
                   // Segundo Convertir a DWORD y hacer SWAP para que el KRC lo lea correctamente
                   #moveCodeKuka := SWAP(UINT_TO_WORD(#code_int));
                   // "moveCodeKuka" := SWAP(UINT_TO_WORD(#code_int));

                   // Dispara GO (flanco por nivel)
                   "goTrigger" := NOT "goTrigger";     // Dispara pedido

                   // Marca estado/ack interno
                   #PlcStatusExecAccepted := TRUE;
                   #PlcStatusExecBusy := TRUE;
                   #PlcStatusExecDone := FALSE;

                   #lastSeq := #KukaControlCmdSeq;          // <-- memoriza!
                   #lastCode := #code_int;             // memoriza qué comando es (para actualizar activos en DONE)

                   #state := 20;                    // BUSY


       END_IF;

   20: // BUSY

       #PlcStatusExecBusy := TRUE;

       #code_int := #KukaControlCmdCode;

       // CANCEL pedido en BUSY → avisar al KRC y ACK de la ORDEN ACTIVA
       IF #code_int = 903 THEN
           "cancelGo" := TRUE;
       END_IF;

       IF ("rbDone" = "goTrigger") THEN
           // Fin confirmado por KUKA

           #PlcStatusExecDone := TRUE;
           #PlcStatusExecBusy := FALSE;
           #PlcStatusExecAccepted := FALSE;
           // ACK de la orden completada
           #PlcStatusExecAckSeq := #lastSeq;

           #state := 0;                         // vuelve a IDLE

       END_IF;

   30: // DONE
       // limpiar y volver a IDLE
       #state := 0;


   END_CASE;
END_REGION
END_FUNCTION_BLOCK

// folder: 20. Robot Services/RobotPos

FUNCTION_BLOCK "TcpPoseDecoderLe32"   // FB4, LAD
{ S7_Optimized_Access := 'TRUE' }
VERSION : 0.1
// Decodifica con SWAP, convierte a DINT y escala.
   VAR_INPUT
      xIniRawLe : DWord;
      yIniRawLe : DWord;
      zIniRawLe : DWord;
      e1IniRawLe : DWord;
      xFinRawLe : DWord;
      yFinRawLe : DWord;
      zFinRawLe : DWord;
      e1FinRawLe : DWord;
      ToolActiveRawByte : Byte;
      BaseActiveRawByte : Byte;
   END_VAR
   VAR_OUTPUT
      tcpPosIniX_mm : LReal;
      tcpPosIniY_mm : LReal;
      tcpPosIniZ_mm : LReal;
      e1PosIni_mm : LReal;
      tcpPosFinX_mm : LReal;
      tcpPosFinY_mm : LReal;
      tcpPosFinZ_mm : LReal;
      e1PosFin_mm : LReal;
      toolActiveId : UDInt;
      baseActiveId : UDInt;
   END_VAR
   VAR_TEMP
      xIniDint : DInt;
      yIniDint : DInt;
      zIniDint : DInt;
      aDint : DInt;
      bDint : DInt;
      cDint : DInt;
      e1IniDint : DInt;
      xFinDint : DInt;
      yFinDint : DInt;
      zFinDint : DInt;
      e1FinDint : DInt;
   END_VAR
BEGIN

REGION Network 1 (SCL): // 1) Endianness: ABCD -> DCBA
   #xIniDint := DWORD_TO_DINT(SWAP(#xIniRawLe));
   #yIniDint := DWORD_TO_DINT(SWAP(#yIniRawLe));
   #zIniDint := DWORD_TO_DINT(SWAP(#zIniRawLe));

   #e1IniDint := DWORD_TO_DINT(SWAP(#e1IniRawLe));

   #xFinDint := DWORD_TO_DINT(SWAP(#xFinRawLe));
   #yFinDint := DWORD_TO_DINT(SWAP(#yFinRawLe));
   #zFinDint := DWORD_TO_DINT(SWAP(#zFinRawLe));
   #e1FinDint := DWORD_TO_DINT(SWAP(#e1FinRawLe));
END_REGION

REGION Network 2 (SCL): // 2) Escala fixed-point: µm->mm, mdeg->deg
   #tcpPosIniX_mm := DINT_TO_LREAL(#xIniDint) / 1000.0;
   #tcpPosIniY_mm := DINT_TO_LREAL(#yIniDint) / 1000.0;
   #tcpPosIniZ_mm := DINT_TO_LREAL(#zIniDint) / 1000.0;

   #e1PosIni_mm := DINT_TO_LREAL(#e1IniDint) / 1000.0;  // mm o deg según tu E1

   #tcpPosFinX_mm := DINT_TO_LREAL(#xFinDint) / 1000.0;
   #tcpPosFinY_mm := DINT_TO_LREAL(#yFinDint) / 1000.0;
   #tcpPosFinZ_mm := DINT_TO_LREAL(#zFinDint) / 1000.0;
   #e1PosFin_mm := DINT_TO_LREAL(#e1FinDint) / 1000.0;  // mm o deg según tu E1

   #toolActiveId := #ToolActiveRawByte;
   #baseActiveId := #BaseActiveRawByte;
END_REGION
END_FUNCTION_BLOCK

// folder: 20. Robot Services/Tooling & Parking

FUNCTION_BLOCK "ToolChange"   // FB6, LAD
TITLE = FB: ManageTed009Station
{ S7_Optimized_Access := 'TRUE' }
VERSION : 0.1
// //  - KUKA manda órdenes (kukaCmd*)
// //  - El FB acciona bobinas de la docking (dockValve*On)
// //  - El FB publica ecos/estados para el KUKA (kukaFeedback*)
// //  - V2 (Unlock) puede mantenerse automática con útil aparcado
// //    (AutoUnlockWhenToolPresent = TRUE) [REF: estándar automático]. 
// //    Con útil ausente, no se activa para evitar soplado innecesario.
// //  - Tapa: FSM con interlock de zona segura y timeouts simétricos.
// //  - Diagnóstico: diagStep/diagFault/diagFaultCode.
// //
// //  Referencias (ver manual Stäubli TED009):
// //    • Sequence plan y sondeo ~20 ms durante conectar/desconectar. 
// //    • +21 mm: E2=0 ∧ E3=1 ∧ D1=0 antes de acoplar. 
// //    • z=0: bloquear retirando V2 y esperar E2=1 ∧ D1=1 (+E1=1). 
// //    • Retiradas +10/+70 y +25/>29 (comentadas para el programa del robot).
   VAR_INPUT
      kukaCmdOpenCover : Bool;
      kukaCmdCloseCover : Bool;
      kukaCmdUnlockMps : Bool;
      kukaCmdSafeForChange : Bool;
      dockSensorToolInPosition : Bool;   // E6
      dockSensorCoverClosed : Bool;   // E4
      dockSensorCoverOpen : Bool;   // E5
      robotSensorMpsUnlocked : Bool;   // E3
      robotSensorMpsLocked : Bool;   // E2
      robotSensorMpsCoupled : Bool;   // E1
      robotSensorMpsCtrlAirPressureOk : Bool;   // D1
      resetFault : Bool;
   END_VAR
   VAR_OUTPUT
      dockValveCoverOpenOn : Bool;   // bobina abrir tapa
      dockValveCoverCloseOn : Bool;   // bobina cerrar tapa
      dockValveV2UnlockOn : Bool;   // V2: aire de desbloqueo hacia módulo del robot
      MpsValveV1B12S4_ON : Bool;
      kukaFeedbackDockCoverOpen : Bool;
      kukaFeedbackDockCoverClosed : Bool;
      kukaFeedbackRobotMpsUnlocked : Bool;
      kukaFeedbackRobotMpsLocked : Bool;
      kukaFeedbackRobotMpsCoupled : Bool;
      kukaFeedbackMpsCtrlAirPressureOk : Bool;
      kukaFeedbackDockToolInPosition : Bool;
      diagStep : Int;
      diagFault : Bool;
      diagFaultCode : Int;
   END_VAR
   VAR
      "step" : Int;
      fault : Bool;
      faultCode : Int;
      AutoUnlockWhenToolPresent : Bool := true;   // // modo auto
      coverTimeout : Time := T#8S;   // // timeout de tapa (abrir/cerrar)
      unlockTimeout : Time := T#2S;   // // timeout de UNLOCK (E3=1 & D1=0)
      unlockReq : Bool;
      unlockReqEnabled : Bool;
      tempCoverOpen : TON_TIME;
      tempCoverClose : TON_TIME;
      tempUnlock : TON_TIME;
      autoUnlockEligible : Bool;
   END_VAR
   VAR CONSTANT
      StateIdle : Int := 0;
      StateOpening : Int := 10;
      StateOpen : Int := 11;
      StateClosing : Int := 20;
      StateClosed : Int := 21;
      FaultNone : Int;
      FaultOpenTimeout : Int := 101;
      FaultCloseTimeout : Int := 102;
      FaultUnlockTimeout : Int := 201;
      FaultInterlock : Int := 301;
   END_VAR
BEGIN

REGION Network 1 (SCL): Lógica de tapa + V2 (Unlock) de la docking
   // --- Feedbacks de estados al robot (eco directo de sensores físicos)
   #kukaFeedbackDockToolInPosition := #dockSensorToolInPosition; // E6 - herramienta en docking station
   #kukaFeedbackDockCoverOpen := #dockSensorCoverOpen;         // E4 - tapa abierta
   #kukaFeedbackDockCoverClosed := #dockSensorCoverClosed;     // E5 - tapa cerrada
   #kukaFeedbackRobotMpsUnlocked := #robotSensorMpsUnlocked;  // E3 - MPS desbloqueado (robot side)
   #kukaFeedbackRobotMpsLocked := #robotSensorMpsLocked;     // E2 - MPS bloqueado (robot side
   #kukaFeedbackRobotMpsCoupled := #robotSensorMpsCoupled;        // E1 - MPS acoplado  (robot side) 
   #kukaFeedbackMpsCtrlAirPressureOk := #robotSensorMpsCtrlAirPressureOk;  // D1 -presostato módulo aire control (robot)
   // ---- Reset de fallos/estado -------------------------------------------
   // Permite reconocer fallos desde HMI/Robot. Pone las salidas a 0 y la FSM (flow state machine)
   // Deja el FB en reposo (IDLE), corta bobinas y reinicia tempor TONs.
   // 
   IF #resetFault THEN
       #fault := FALSE;
       #faultCode := #FaultNone;
       #step := #StateIdle;

       #dockValveCoverOpenOn := FALSE;
       #dockValveCoverCloseOn := FALSE;
       #dockValveV2UnlockOn := FALSE;

       // Reset explícito de TON: IN=FALSE + PT definido
       #tempCoverOpen(IN := FALSE,
                      PT := #coverTimeout);
       #tempCoverClose(IN := FALSE,
                       PT := #coverTimeout);
       #tempUnlock(IN := FALSE,
                   PT := #unlockTimeout);
   END_IF;

   // ================= LÓGICA DE TAPA (máquina de estados) =================
   // Interlock básico: no se permite accionar tapa si el robot no confirma zona segura
   // (manual: abrir/cerrar solo fuera del barrido).
   CASE #step OF

       #StateIdle: // IDLE
           // Reposo ( tapa sin accionar); evaluar órdenes de KUKA.
           #dockValveCoverOpenOn := FALSE;
           #dockValveCoverCloseOn := FALSE;

           IF #kukaCmdSafeForChange THEN
               // Abrir si lo pide el robot y aún no está abierta
               IF (#kukaCmdOpenCover AND NOT #dockSensorCoverOpen) THEN
                   #step := #StateOpening;
               END_IF;
               // Cerrar si lo pide el robot y aún no está cerrada
               IF (#kukaCmdCloseCover AND NOT #dockSensorCoverClosed) THEN
                   #step := #StateClosing;
               END_IF;
           ELSIF (#kukaCmdOpenCover OR #kukaCmdCloseCover) THEN
               // Petición sin zona segura -> fallo de interlock
               #fault := TRUE;
               #faultCode := #FaultInterlock; // robot no garantiza zona segura
           END_IF;

       #StateOpening:  // Abrir tapa
           #dockValveCoverOpenOn := TRUE;
           #dockValveCoverCloseOn := FALSE;

           // Timeout de apertura: si no llega "tapa abierta" dentro de coverTimeout -> fallo.
           // coverTimeout debe ser > 3 s (tiempo típico de maniobra)
           #tempCoverOpen(IN := NOT #dockSensorCoverOpen,
                          PT := #coverTimeout);

           IF (#dockSensorCoverOpen AND NOT #dockSensorCoverClosed) THEN
               #tempCoverOpen(IN := FALSE,
                              PT := #coverTimeout);
               #step := #StateOpen;
           ELSIF #tempCoverOpen.Q THEN
               #fault := TRUE;
               #faultCode := #FaultOpenTimeout;
               #dockValveCoverOpenOn := FALSE;
               #step := #StateIdle;
           END_IF;

       #StateOpen: // Tapa abierta (estable)
           #dockValveCoverOpenOn := FALSE;
           #dockValveCoverCloseOn := FALSE;

           IF (#kukaCmdSafeForChange AND #kukaCmdCloseCover) THEN
               #step := #StateClosing;
           END_IF;


       #StateClosing: // Cerrar tapa
           #dockValveCoverOpenOn := FALSE;
           #dockValveCoverCloseOn := TRUE;

           // Timeout de cierre: si no llega "tapa cerrada" dentro de coverTimeout -> fallo.
           #tempCoverClose(IN := NOT #dockSensorCoverClosed,
                           PT := #coverTimeout);

           IF (#dockSensorCoverClosed AND NOT #dockSensorCoverOpen) THEN
               #tempCoverClose(IN := FALSE,
                               PT := #coverTimeout);
               #step := #StateClosed;
           ELSIF #tempCoverClose.Q THEN
               #fault := TRUE;
               #faultCode := #FaultCloseTimeout;
               #dockValveCoverCloseOn := FALSE;
               #step := #StateIdle;
           END_IF;

       #StateClosed: // Tapa cerrada (estable)
           #dockValveCoverOpenOn := FALSE;
           #dockValveCoverCloseOn := FALSE;

           IF (#kukaCmdSafeForChange AND #kukaCmdOpenCover) THEN
               #step := #StateOpening;
           END_IF;

       ELSE
           #step := #StateIdle;
   END_CASE;

   // Exclusión mutua de bobinas de tapa (seguridad por si alguna rama dejó ambas a 1)
   IF #dockValveCoverOpenOn THEN
       #dockValveCoverCloseOn := FALSE;
   END_IF;
   IF #dockValveCoverCloseOn THEN
       #dockValveCoverOpenOn := FALSE;
   END_IF;



   // -------- Arbitraje de V2 (UNLOCK) — sin auto-unlock --------
   #autoUnlockEligible := FALSE;   // DEPRECATED: ya no se usa

   //Cuando el robot va al punto de acople hace antes kukaCmdUnlockMpsYugo = TRUE

   //  solo por orden KUKA 
   #dockValveV2UnlockOn := #kukaCmdUnlockMps;

   IF #robotSensorMpsLocked THEN
       #MpsValveV1B12S4_ON := TRUE;
   END_IF;


   // Supervisión del estado desbloqueado (E3=1 y D1=0 en tiempo):
   #tempUnlock(
               IN := (#dockValveV2UnlockOn
               AND NOT (#robotSensorMpsUnlocked
               AND NOT #robotSensorMpsCtrlAirPressureOk)),
               PT := #unlockTimeout
   );
   IF NOT #dockValveV2UnlockOn THEN
       // reset explícito del TON cuando ya no se pide V2
       #tempUnlock(IN := FALSE,
                   PT := #unlockTimeout);
   END_IF;

   // -------------------- DIAGNÓSTICO PUBLICADO ----------------------------
   #diagStep := #step; // StateIdle/Opening/Open/Closing/Closed
   #diagFault := #fault;
   #diagFaultCode := #faultCode;
END_REGION
END_FUNCTION_BLOCK

FUNCTION_BLOCK "MpsDockingStation"   // FB9, LAD
{ S7_Optimized_Access := 'TRUE' }
VERSION : 0.1
BEGIN

REGION Network 1: Identificador de Herramienta
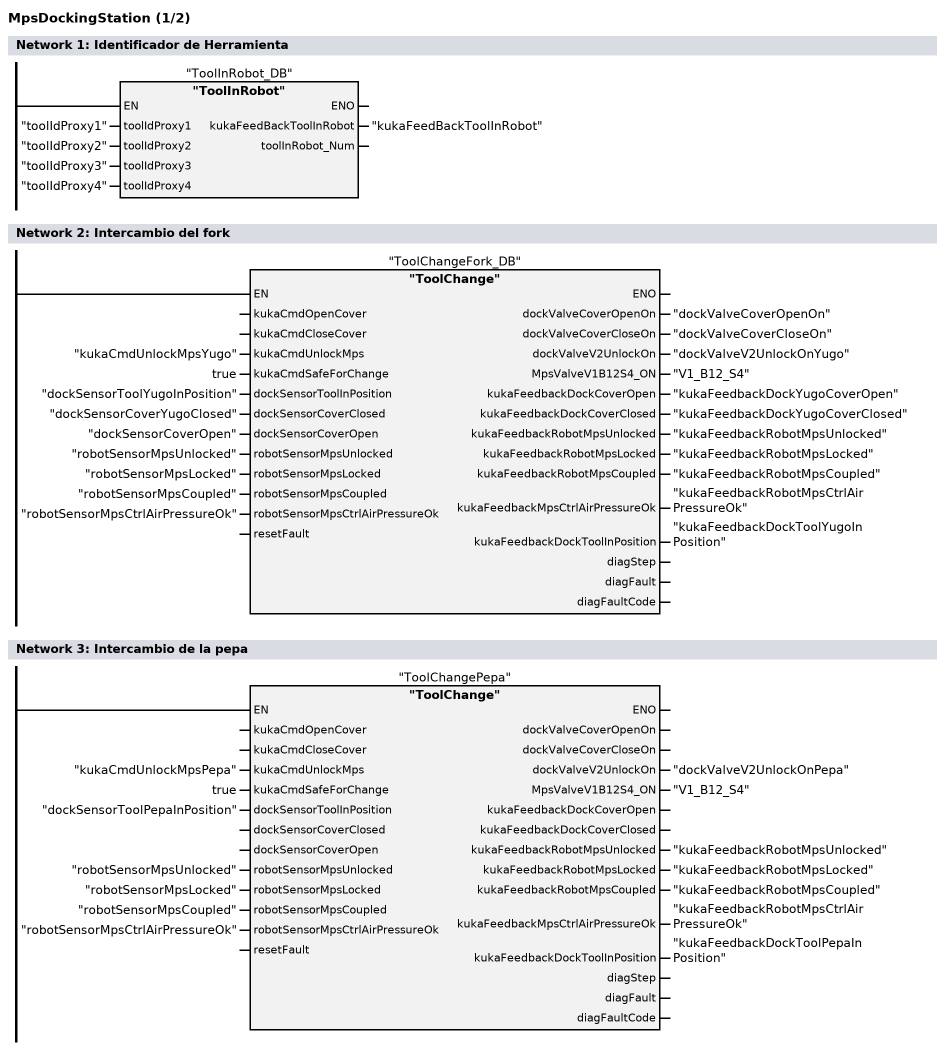
   RUNG wire#powerrail
      "ToolInRobot_DB"(toolIdProxy1 := "toolIdProxy1", toolIdProxy2 := "toolIdProxy2", toolIdProxy3 := "toolIdProxy3", toolIdProxy4 := "toolIdProxy4", kukaFeedBackToolInRobot => "kukaFeedBackToolInRobot", toolInRobot_Num =>)
   END_RUNG
   // the same network as SCL:
   "ToolInRobot_DB"(toolIdProxy1 := "toolIdProxy1",   // "ToolInRobot"
                    toolIdProxy2 := "toolIdProxy2",
                    toolIdProxy3 := "toolIdProxy3",
                    toolIdProxy4 := "toolIdProxy4",
                    kukaFeedBackToolInRobot => "kukaFeedBackToolInRobot");
END_REGION

REGION Network 2: Intercambio del fork
   RUNG wire#powerrail
      "ToolChangeFork_DB"(kukaCmdOpenCover :=, kukaCmdCloseCover :=, kukaCmdUnlockMps := "kukaCmdUnlockMpsYugo", kukaCmdSafeForChange := true, dockSensorToolInPosition := "dockSensorToolYugoInPosition", dockSensorCoverClosed := "dockSensorCoverYugoClosed", dockSensorCoverOpen := "dockSensorCoverOpen", robotSensorMpsUnlocked := "robotSensorMpsUnlocked", robotSensorMpsLocked := "robotSensorMpsLocked", robotSensorMpsCoupled := "robotSensorMpsCoupled", robotSensorMpsCtrlAirPressureOk := "robotSensorMpsCtrlAirPressureOk", resetFault :=, dockValveCoverOpenOn => "dockValveCoverOpenOn", dockValveCoverCloseOn => "dockValveCoverCloseOn", dockValveV2UnlockOn => "dockValveV2UnlockOnYugo", MpsValveV1B12S4_ON => "V1_B12_S4", kukaFeedbackDockCoverOpen => "kukaFeedbackDockYugoCoverOpen", kukaFeedbackDockCoverClosed => "kukaFeedbackDockYugoCoverClosed", kukaFeedbackRobotMpsUnlocked => "kukaFeedbackRobotMpsUnlocked", kukaFeedbackRobotMpsLocked => "kukaFeedbackRobotMpsLocked", kukaFeedbackRobotMpsCoupled => "kukaFeedbackRobotMpsCoupled", kukaFeedbackMpsCtrlAirPressureOk => "kukaFeedbackRobotMpsCtrlAirPressureOk", kukaFeedbackDockToolInPosition => "kukaFeedbackDockToolYugoInPosition", diagStep =>, diagFault =>, diagFaultCode =>)
   END_RUNG
   // the same network as SCL:
   "ToolChangeFork_DB"(kukaCmdUnlockMps := "kukaCmdUnlockMpsYugo",   // "ToolChange"
                       kukaCmdSafeForChange := true,
                       dockSensorToolInPosition := "dockSensorToolYugoInPosition",
                       dockSensorCoverClosed := "dockSensorCoverYugoClosed",
                       dockSensorCoverOpen := "dockSensorCoverOpen",
                       robotSensorMpsUnlocked := "robotSensorMpsUnlocked",
                       robotSensorMpsLocked := "robotSensorMpsLocked",
                       robotSensorMpsCoupled := "robotSensorMpsCoupled",
                       robotSensorMpsCtrlAirPressureOk := "robotSensorMpsCtrlAirPressureOk",
                       dockValveCoverOpenOn => "dockValveCoverOpenOn",
                       dockValveCoverCloseOn => "dockValveCoverCloseOn",
                       dockValveV2UnlockOn => "dockValveV2UnlockOnYugo",
                       MpsValveV1B12S4_ON => "V1_B12_S4",
                       kukaFeedbackDockCoverOpen => "kukaFeedbackDockYugoCoverOpen",
                       kukaFeedbackDockCoverClosed => "kukaFeedbackDockYugoCoverClosed",
                       kukaFeedbackRobotMpsUnlocked => "kukaFeedbackRobotMpsUnlocked",
                       kukaFeedbackRobotMpsLocked => "kukaFeedbackRobotMpsLocked",
                       kukaFeedbackRobotMpsCoupled => "kukaFeedbackRobotMpsCoupled",
                       kukaFeedbackMpsCtrlAirPressureOk => "kukaFeedbackRobotMpsCtrlAirPressureOk",
                       kukaFeedbackDockToolInPosition => "kukaFeedbackDockToolYugoInPosition");
END_REGION

REGION Network 3: Intercambio de la pepa
   RUNG wire#powerrail
      "ToolChangePepa"(kukaCmdOpenCover :=, kukaCmdCloseCover :=, kukaCmdUnlockMps := "kukaCmdUnlockMpsPepa", kukaCmdSafeForChange := true, dockSensorToolInPosition := "dockSensorToolPepaInPosition", dockSensorCoverClosed :=, dockSensorCoverOpen :=, robotSensorMpsUnlocked := "robotSensorMpsUnlocked", robotSensorMpsLocked := "robotSensorMpsLocked", robotSensorMpsCoupled := "robotSensorMpsCoupled", robotSensorMpsCtrlAirPressureOk := "robotSensorMpsCtrlAirPressureOk", resetFault :=, dockValveCoverOpenOn =>, dockValveCoverCloseOn =>, dockValveV2UnlockOn => "dockValveV2UnlockOnPepa", MpsValveV1B12S4_ON => "V1_B12_S4", kukaFeedbackDockCoverOpen =>, kukaFeedbackDockCoverClosed =>, kukaFeedbackRobotMpsUnlocked => "kukaFeedbackRobotMpsUnlocked", kukaFeedbackRobotMpsLocked => "kukaFeedbackRobotMpsLocked", kukaFeedbackRobotMpsCoupled => "kukaFeedbackRobotMpsCoupled", kukaFeedbackMpsCtrlAirPressureOk => "kukaFeedbackRobotMpsCtrlAirPressureOk", kukaFeedbackDockToolInPosition => "kukaFeedbackDockToolPepaInPosition", diagStep =>, diagFault =>, diagFaultCode =>)
   END_RUNG
   // the same network as SCL:
   "ToolChangePepa"(kukaCmdUnlockMps := "kukaCmdUnlockMpsPepa",   // "ToolChange"
                    kukaCmdSafeForChange := true,
                    dockSensorToolInPosition := "dockSensorToolPepaInPosition",
                    robotSensorMpsUnlocked := "robotSensorMpsUnlocked",
                    robotSensorMpsLocked := "robotSensorMpsLocked",
                    robotSensorMpsCoupled := "robotSensorMpsCoupled",
                    robotSensorMpsCtrlAirPressureOk := "robotSensorMpsCtrlAirPressureOk",
                    dockValveV2UnlockOn => "dockValveV2UnlockOnPepa",
                    MpsValveV1B12S4_ON => "V1_B12_S4",
                    kukaFeedbackRobotMpsUnlocked => "kukaFeedbackRobotMpsUnlocked",
                    kukaFeedbackRobotMpsLocked => "kukaFeedbackRobotMpsLocked",
                    kukaFeedbackRobotMpsCoupled => "kukaFeedbackRobotMpsCoupled",
                    kukaFeedbackMpsCtrlAirPressureOk => "kukaFeedbackRobotMpsCtrlAirPressureOk",
                    kukaFeedbackDockToolInPosition => "kukaFeedbackDockToolPepaInPosition");
END_REGION

REGION Network 4: Intercambio de la heramienta de Inmersion - Pole
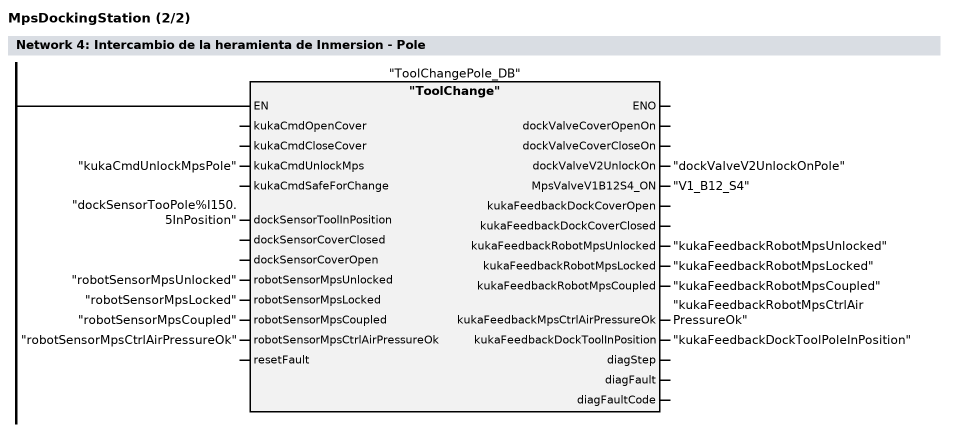
   RUNG wire#powerrail
      "ToolChangePole_DB"(kukaCmdOpenCover :=, kukaCmdCloseCover :=, kukaCmdUnlockMps := "kukaCmdUnlockMpsPole", kukaCmdSafeForChange :=, dockSensorToolInPosition := "dockSensorTooPole%I150.5InPosition", dockSensorCoverClosed :=, dockSensorCoverOpen :=, robotSensorMpsUnlocked := "robotSensorMpsUnlocked", robotSensorMpsLocked := "robotSensorMpsLocked", robotSensorMpsCoupled := "robotSensorMpsCoupled", robotSensorMpsCtrlAirPressureOk := "robotSensorMpsCtrlAirPressureOk", resetFault :=, dockValveCoverOpenOn =>, dockValveCoverCloseOn =>, dockValveV2UnlockOn => "dockValveV2UnlockOnPole", MpsValveV1B12S4_ON => "V1_B12_S4", kukaFeedbackDockCoverOpen =>, kukaFeedbackDockCoverClosed =>, kukaFeedbackRobotMpsUnlocked => "kukaFeedbackRobotMpsUnlocked", kukaFeedbackRobotMpsLocked => "kukaFeedbackRobotMpsLocked", kukaFeedbackRobotMpsCoupled => "kukaFeedbackRobotMpsCoupled", kukaFeedbackMpsCtrlAirPressureOk => "kukaFeedbackRobotMpsCtrlAirPressureOk", kukaFeedbackDockToolInPosition => "kukaFeedbackDockToolPoleInPosition", diagStep =>, diagFault =>, diagFaultCode =>)
   END_RUNG
   // the same network as SCL:
   "ToolChangePole_DB"(kukaCmdUnlockMps := "kukaCmdUnlockMpsPole",   // "ToolChange"
                       dockSensorToolInPosition := "dockSensorTooPole%I150.5InPosition",
                       robotSensorMpsUnlocked := "robotSensorMpsUnlocked",
                       robotSensorMpsLocked := "robotSensorMpsLocked",
                       robotSensorMpsCoupled := "robotSensorMpsCoupled",
                       robotSensorMpsCtrlAirPressureOk := "robotSensorMpsCtrlAirPressureOk",
                       dockValveV2UnlockOn => "dockValveV2UnlockOnPole",
                       MpsValveV1B12S4_ON => "V1_B12_S4",
                       kukaFeedbackRobotMpsUnlocked => "kukaFeedbackRobotMpsUnlocked",
                       kukaFeedbackRobotMpsLocked => "kukaFeedbackRobotMpsLocked",
                       kukaFeedbackRobotMpsCoupled => "kukaFeedbackRobotMpsCoupled",
                       kukaFeedbackMpsCtrlAirPressureOk => "kukaFeedbackRobotMpsCtrlAirPressureOk",
                       kukaFeedbackDockToolInPosition => "kukaFeedbackDockToolPoleInPosition");
END_REGION
END_FUNCTION_BLOCK

FUNCTION_BLOCK "ToolInRobot"   // FB15, LAD
{ S7_Optimized_Access := 'TRUE' }
VERSION : 0.1
   VAR_INPUT
      toolIdProxy1 : Bool;
      toolIdProxy2 : Bool;
      toolIdProxy3 : Bool;
      toolIdProxy4 : Bool;
   END_VAR
   VAR_OUTPUT
      kukaFeedBackToolInRobot : Word;
      toolInRobot_Num : UInt;
   END_VAR
   VAR_TEMP
      mask : Byte;
   END_VAR
BEGIN

REGION Network 1 (SCL)

   #mask := 0;
   IF #toolIdProxy1 THEN
       #mask := #mask + 1;
   END_IF;   // bit0
   IF #toolIdProxy2 THEN
       #mask := #mask + 2;
   END_IF;   // bit1
   IF #toolIdProxy3 THEN
       #mask := #mask + 4;
   END_IF;   // bit2
   IF #toolIdProxy4 THEN
       #mask := #mask + 8;
   END_IF;   // bit3

   //Stand 1 - Tool 1 - Fork 
   //Stand 2 - Tool 2 - Pepa
   //Stand 3 - TOOL 3 - Marker
   //Stand 4 - Tool 4 - Gocator
   //Stand 5 - Tool 5 - Pole
   //Falta ajustar los sensores para que generen esas combinaciones.

   CASE #mask OF

       0:
           #toolInRobot_Num := 0;   // sin herramienta
           #kukaFeedBackToolInRobot := SWAP(UINT_TO_WORD(#toolInRobot_Num));
       1:
           #toolInRobot_Num := 2;   // PEPA
           #kukaFeedBackToolInRobot := SWAP(UINT_TO_WORD(#toolInRobot_Num));
       2:
           #toolInRobot_Num := 5;   // pole
           #kukaFeedBackToolInRobot := SWAP(UINT_TO_WORD(#toolInRobot_Num));
       3:
           #toolInRobot_Num := 1;   // fork
           #kukaFeedBackToolInRobot := SWAP(UINT_TO_WORD(#toolInRobot_Num));
          // #kukaFeedBackToolInRobot := UINT_TO_WORD(#toolInRobot_Num);  // SIN SWAP
       4:
           #toolInRobot_Num := 4;   // teaching
           #kukaFeedBackToolInRobot := SWAP(UINT_TO_WORD(#toolInRobot_Num));
       5:
           #toolInRobot_Num := 3;   // marker
           #kukaFeedBackToolInRobot := SWAP(UINT_TO_WORD(#toolInRobot_Num));
       ELSE
           #toolInRobot_Num := -1;      // combinación no válida / desconocida
   END_CASE;
END_REGION
END_FUNCTION_BLOCK

// folder: 30. Safety

FUNCTION_BLOCK "MainSafety"   // FB1, F_LAD
{ S7_Optimized_Access := 'TRUE' }
// // Functionality: Monitoring of the protective door position, light curtain and emergency stop
   VAR
      ACK_GL_Instance : ACK_GL;
      instEStopGroup : "EStopGroup";
      instLightCurtainGroup : "LightCurtainGroup";
      instSafetyDoor : "SafetyDoor";
      SafetyRobot_Instance : "SafetyRobot";
   END_VAR
   VAR_TEMP
      tempEStop1Released : Bool;
      tempEStop2Released : Bool;
      tempEStop3Released : Bool;
      tempEStop4Released : Bool;
      tempEStop5Released : Bool;
      tempEStop6Released : Bool;
      tempEStop7Released : Bool;
      tempEStop8Released : Bool;
      tempEStopAllReleased : Bool;
      tempEStopReleasedActuator : Bool;
      tempEStopAckReq : Bool;
      tempLc1Free : Bool;
      tempLc2Free : Bool;
      tempLc3Free : Bool;
      tempLc4Free : Bool;
      tempLc5Free : Bool;
      tempLc6Free : Bool;
      tempLcAllFree : Bool;
      tempLcAccessGrantedZ1 : Bool;
      tempLcAccessGrantedZ2 : Bool;
      tempLcAccessGrantedZ3 : Bool;
   END_VAR
BEGIN

REGION Network 1: Emergency stop
   // When the emergency stop is pressed, the actuator becomes safe switched off.
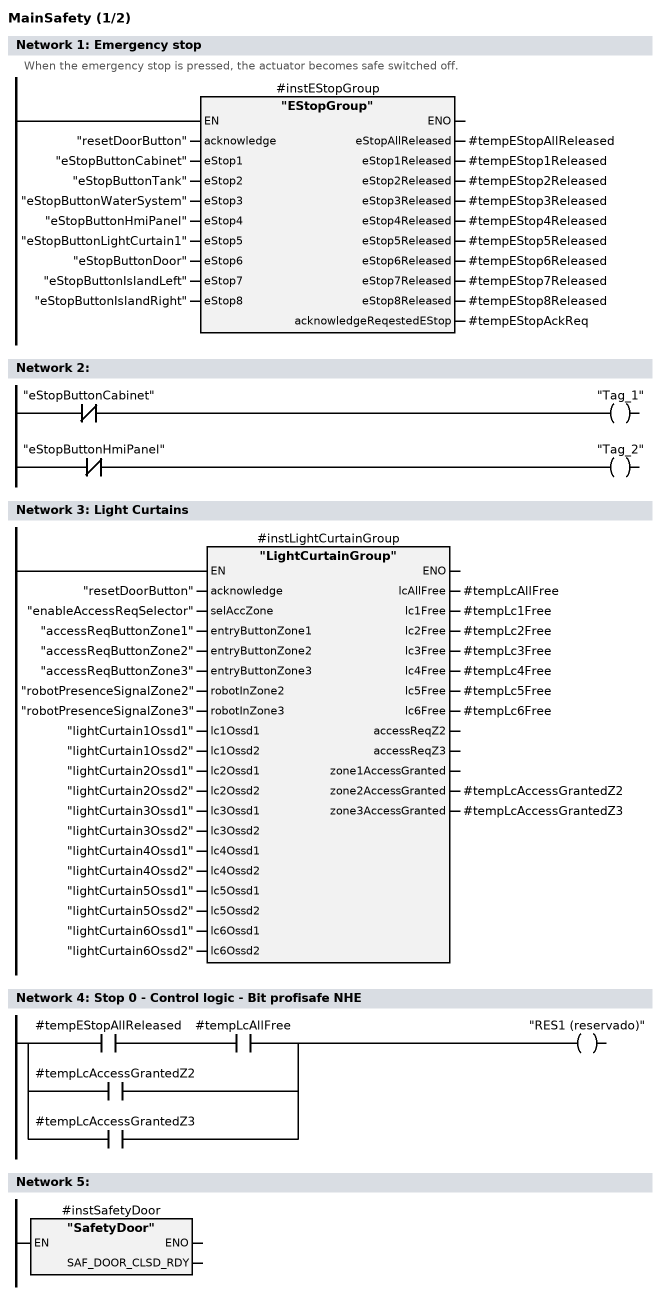
   RUNG wire#powerrail
      #instEStopGroup(acknowledge := "resetDoorButton", eStop1 := "eStopButtonCabinet", eStop2 := "eStopButtonTank", eStop3 := "eStopButtonWaterSystem", eStop4 := "eStopButtonHmiPanel", eStop5 := "eStopButtonLightCurtain1", eStop6 := "eStopButtonDoor", eStop7 := "eStopButtonIslandLeft", eStop8 := "eStopButtonIslandRight", eStopAllReleased => #tempEStopAllReleased, eStop1Released => #tempEStop1Released, eStop2Released => #tempEStop2Released, eStop3Released => #tempEStop3Released, eStop4Released => #tempEStop4Released, eStop5Released => #tempEStop5Released, eStop6Released => #tempEStop6Released, eStop7Released => #tempEStop7Released, eStop8Released => #tempEStop8Released, acknowledgeReqestedEStop => #tempEStopAckReq)
   END_RUNG
   // the same network as SCL:
   #instEStopGroup(acknowledge := "resetDoorButton",   // "EStopGroup"
                   eStop1 := "eStopButtonCabinet",
                   eStop2 := "eStopButtonTank",
                   eStop3 := "eStopButtonWaterSystem",
                   eStop4 := "eStopButtonHmiPanel",
                   eStop5 := "eStopButtonLightCurtain1",
                   eStop6 := "eStopButtonDoor",
                   eStop7 := "eStopButtonIslandLeft",
                   eStop8 := "eStopButtonIslandRight",
                   eStopAllReleased => #tempEStopAllReleased,
                   eStop1Released => #tempEStop1Released,
                   eStop2Released => #tempEStop2Released,
                   eStop3Released => #tempEStop3Released,
                   eStop4Released => #tempEStop4Released,
                   eStop5Released => #tempEStop5Released,
                   eStop6Released => #tempEStop6Released,
                   eStop7Released => #tempEStop7Released,
                   eStop8Released => #tempEStop8Released,
                   acknowledgeReqestedEStop => #tempEStopAckReq);
END_REGION

REGION Network 2
   RUNG wire#powerrail
      I_Contact( "eStopButtonCabinet" )
      Coil( "Tag_1" )
   END_RUNG
   RUNG wire#powerrail
      I_Contact( "eStopButtonHmiPanel" )
      Coil( "Tag_2" )
   END_RUNG
   // the same network as SCL:
   "Tag_1" := NOT "eStopButtonCabinet";
   "Tag_2" := NOT "eStopButtonHmiPanel";
END_REGION

REGION Network 3: Light Curtains
   RUNG wire#powerrail
      #instLightCurtainGroup(acknowledge := "resetDoorButton", selAccZone := "enableAccessReqSelector", entryButtonZone1 := "accessReqButtonZone1", entryButtonZone2 := "accessReqButtonZone2", entryButtonZone3 := "accessReqButtonZone3", robotInZone2 := "robotPresenceSignalZone2", robotInZone3 := "robotPresenceSignalZone3", lc1Ossd1 := "lightCurtain1Ossd1", lc1Ossd2 := "lightCurtain1Ossd2", lc2Ossd1 := "lightCurtain2Ossd1", lc2Ossd2 := "lightCurtain2Ossd2", lc3Ossd1 := "lightCurtain3Ossd1", lc3Ossd2 := "lightCurtain3Ossd2", lc4Ossd1 := "lightCurtain4Ossd1", lc4Ossd2 := "lightCurtain4Ossd2", lc5Ossd1 := "lightCurtain5Ossd1", lc5Ossd2 := "lightCurtain5Ossd2", lc6Ossd1 := "lightCurtain6Ossd1", lc6Ossd2 := "lightCurtain6Ossd2", lcAllFree => #tempLcAllFree, lc1Free => #tempLc1Free, lc2Free => #tempLc2Free, lc3Free => #tempLc3Free, lc4Free => #tempLc4Free, lc5Free => #tempLc5Free, lc6Free => #tempLc6Free, accessReqZ2 =>, accessReqZ3 =>, zone1AccessGranted =>, zone2AccessGranted => #tempLcAccessGrantedZ2, zone3AccessGranted => #tempLcAccessGrantedZ3)
   END_RUNG
   // the same network as SCL:
   #instLightCurtainGroup(acknowledge := "resetDoorButton",   // "LightCurtainGroup"
                          selAccZone := "enableAccessReqSelector",
                          entryButtonZone1 := "accessReqButtonZone1",
                          entryButtonZone2 := "accessReqButtonZone2",
                          entryButtonZone3 := "accessReqButtonZone3",
                          robotInZone2 := "robotPresenceSignalZone2",
                          robotInZone3 := "robotPresenceSignalZone3",
                          lc1Ossd1 := "lightCurtain1Ossd1",
                          lc1Ossd2 := "lightCurtain1Ossd2",
                          lc2Ossd1 := "lightCurtain2Ossd1",
                          lc2Ossd2 := "lightCurtain2Ossd2",
                          lc3Ossd1 := "lightCurtain3Ossd1",
                          lc3Ossd2 := "lightCurtain3Ossd2",
                          lc4Ossd1 := "lightCurtain4Ossd1",
                          lc4Ossd2 := "lightCurtain4Ossd2",
                          lc5Ossd1 := "lightCurtain5Ossd1",
                          lc5Ossd2 := "lightCurtain5Ossd2",
                          lc6Ossd1 := "lightCurtain6Ossd1",
                          lc6Ossd2 := "lightCurtain6Ossd2",
                          lcAllFree => #tempLcAllFree,
                          lc1Free => #tempLc1Free,
                          lc2Free => #tempLc2Free,
                          lc3Free => #tempLc3Free,
                          lc4Free => #tempLc4Free,
                          lc5Free => #tempLc5Free,
                          lc6Free => #tempLc6Free,
                          zone2AccessGranted => #tempLcAccessGrantedZ2,
                          zone3AccessGranted => #tempLcAccessGrantedZ3);
END_REGION

REGION Network 4: Stop 0 - Control logic - Bit profisafe NHE
   RUNG wire#powerrail
      Contact( #tempEStopAllReleased )
      Contact( #tempLcAllFree )
      wire#w1
      Coil( "RES1 (reservado)" )
   END_RUNG
   RUNG wire#powerrail
      Contact( #tempLcAccessGrantedZ2 )
   END_RUNG wire#w1
   RUNG wire#powerrail
      Contact( #tempLcAccessGrantedZ3 )
   END_RUNG wire#w1
   // the same network as SCL:
   "RES1 (reservado)" := (#tempEStopAllReleased AND #tempLcAllFree) OR #tempLcAccessGrantedZ2 OR #tempLcAccessGrantedZ3;
END_REGION

REGION Network 5
   RUNG wire#powerrail
      #instSafetyDoor(SAF_DOOR_CLSD_RDY =>)
   END_RUNG
   // the same network as SCL:
   #instSafetyDoor();   // "SafetyDoor"
END_REGION

REGION Network 6
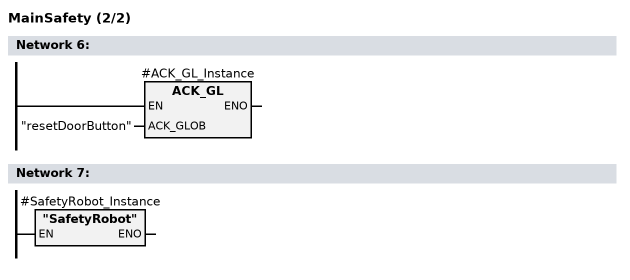
   #ACK_GL_Instance(ACK_GLOB := "resetDoorButton");   // ACK_GL
END_REGION

REGION Network 7
   RUNG wire#powerrail
      #SafetyRobot_Instance()
   END_RUNG
   // the same network as SCL:
   #SafetyRobot_Instance();   // "SafetyRobot"
END_REGION
END_FUNCTION_BLOCK

FUNCTION_BLOCK "SafetyRobot"   // FB3, F_LAD
{ S7_Optimized_Access := 'TRUE' }
VERSION : 0.1
   VAR
      Edge_ACK : Bool;
      mem_ack_trig : Bool;
      ACK_GL_Instance : Bool;
      F_IEC_Timer_Instance_1 : TP;
   END_VAR
   VAR_TEMP   // added for the SCL form of the ladder/FBD networks
      _w1 : Bool;
   END_VAR
BEGIN

REGION Network 1: Reservado (debe ser 1)
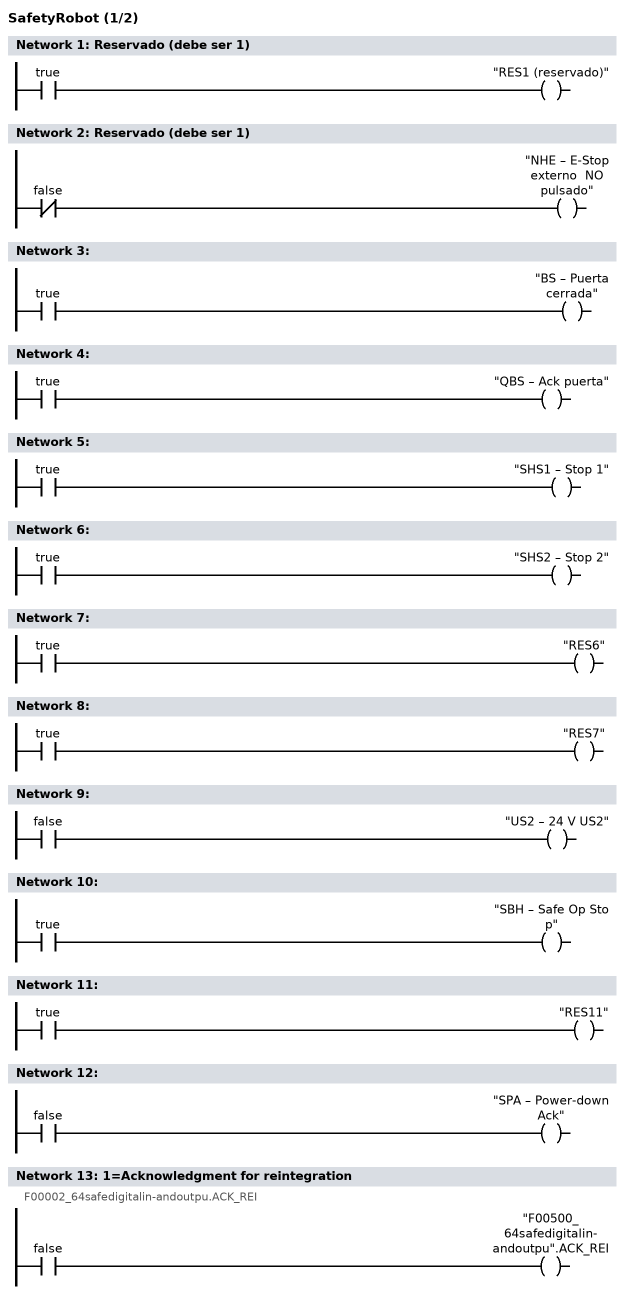
   RUNG wire#powerrail
      Contact( true )
      Coil( "RES1 (reservado)" )
   END_RUNG
   // the same network as SCL:
   "RES1 (reservado)" := true;
END_REGION

REGION Network 2: Reservado (debe ser 1)
   RUNG wire#powerrail
      I_Contact( false )
      Coil( "NHE – E‑Stop externo  NO pulsado" )
   END_RUNG
   // the same network as SCL:
   "NHE – E‑Stop externo  NO pulsado" := NOT false;
END_REGION

REGION Network 3
   RUNG wire#powerrail
      Contact( true )
      Coil( "BS – Puerta cerrada" )
   END_RUNG
   // the same network as SCL:
   "BS – Puerta cerrada" := true;
END_REGION

REGION Network 4
   RUNG wire#powerrail
      Contact( true )
      Coil( "QBS – Ack puerta" )
   END_RUNG
   // the same network as SCL:
   "QBS – Ack puerta" := true;
END_REGION

REGION Network 5
   RUNG wire#powerrail
      Contact( true )
      Coil( "SHS1 – Stop 1" )
   END_RUNG
   // the same network as SCL:
   "SHS1 – Stop 1" := true;
END_REGION

REGION Network 6
   RUNG wire#powerrail
      Contact( true )
      Coil( "SHS2 – Stop 2" )
   END_RUNG
   // the same network as SCL:
   "SHS2 – Stop 2" := true;
END_REGION

REGION Network 7
   RUNG wire#powerrail
      Contact( true )
      Coil( "RES6" )
   END_RUNG
   // the same network as SCL:
   "RES6" := true;
END_REGION

REGION Network 8
   RUNG wire#powerrail
      Contact( true )
      Coil( "RES7" )
   END_RUNG
   // the same network as SCL:
   "RES7" := true;
END_REGION

REGION Network 9
   RUNG wire#powerrail
      Contact( false )
      Coil( "US2 – 24 V US2" )
   END_RUNG
   // the same network as SCL:
   "US2 – 24 V US2" := false;
END_REGION

REGION Network 10
   RUNG wire#powerrail
      Contact( true )
      Coil( "SBH – Safe Op Stop" )
   END_RUNG
   // the same network as SCL:
   "SBH – Safe Op Stop" := true;
END_REGION

REGION Network 11
   RUNG wire#powerrail
      Contact( true )
      Coil( "RES11" )
   END_RUNG
   // the same network as SCL:
   "RES11" := true;
END_REGION

REGION Network 12
   RUNG wire#powerrail
      Contact( false )
      Coil( "SPA – Power‑down Ack" )
   END_RUNG
   // the same network as SCL:
   "SPA – Power‑down Ack" := false;
END_REGION

REGION Network 13: 1=Acknowledgment for reintegration
   // F00002_64safedigitalin-andoutpu.ACK_REI
   RUNG wire#powerrail
      Contact( false )
      Coil( "F00500_64safedigitalin-andoutpu".ACK_REI )
   END_RUNG
   // the same network as SCL:
   "F00500_64safedigitalin-andoutpu".ACK_REI := false;
END_REGION

REGION Network 14: Pulse output
   // - CLK → F00002_…ACK_REQ : Detecta el flanco 0 → 1 que el módulo pone cuando necesita
   // - M → mem_ACK_Trig
   // : reconocimiento. El 1 sólo dura un scan y se guarda internamente en mem_ACK_Trig….
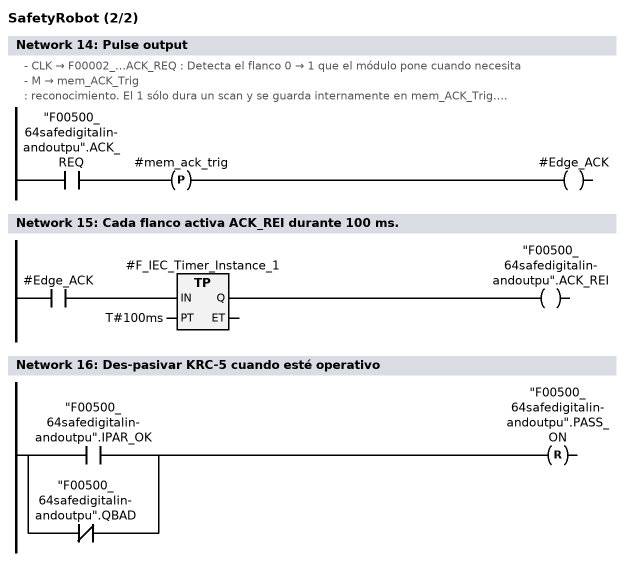
   RUNG wire#powerrail
      Contact( "F00500_64safedigitalin-andoutpu".ACK_REQ )
      P_Trig( #mem_ack_trig )
      Coil( #Edge_ACK )
   END_RUNG
   // the same network as SCL:
   #_w1 := "F00500_64safedigitalin-andoutpu".ACK_REQ AND NOT #mem_ack_trig;   // rising edge
   #mem_ack_trig := "F00500_64safedigitalin-andoutpu".ACK_REQ;
   #Edge_ACK := #_w1;
END_REGION

REGION Network 15: Cada flanco activa ACK_REI durante 100 ms.
   #F_IEC_Timer_Instance_1.TP(IN := #Edge_ACK, PT := T#100ms);
   "F00500_64safedigitalin-andoutpu".ACK_REI := #F_IEC_Timer_Instance_1.Q;
END_REGION

REGION Network 16: Des-pasivar KRC-5 cuando esté operativo
   RUNG wire#powerrail
      Contact( "F00500_64safedigitalin-andoutpu".IPAR_OK )
      wire#w1
      R_Coil( "F00500_64safedigitalin-andoutpu".PASS_ON )
   END_RUNG
   RUNG wire#powerrail
      I_Contact( "F00500_64safedigitalin-andoutpu".QBAD )
   END_RUNG wire#w1
   // the same network as SCL:
   IF "F00500_64safedigitalin-andoutpu".IPAR_OK OR NOT "F00500_64safedigitalin-andoutpu".QBAD THEN
       "F00500_64safedigitalin-andoutpu".PASS_ON := FALSE;
   END_IF;
END_REGION
END_FUNCTION_BLOCK

// folder: 30. Safety/SafetyFunctions

FUNCTION_BLOCK "EStopGroup"   // FB2, F_LAD
{ S7_Optimized_Access := 'TRUE' }